   Button "b_Save" at 1074,510 size 72x64; TextOff 'SAVE'; Authorization "Operate"; PictureOff "SetHD"
      on Click: SetBit("DB_MouldEditor_HMI_uData_sStatusBits_xSafeChanges"); "VBStore_tool"('\Storage Card SD')
      Visibility <- "DB_MouldEditor_HMI_uData_sStatusBits_xValueChanged"
   IOField "I/O field_15" at 673,669 size 77x35; Authorization "Operate"; FormatPattern 9999.99
      ProcessValue <- "DB_MouldEditor_HMI_uData_sSelected_sPS_arFlow{3}"
      Visibility <- "DB704_MH_Value_Mixinghead{0}_AmountComponent"
      ObjectEnable <- "DB_MouldEditor_HMI_uData_sSelected_iCalculation"
      Appearance <- "DB_MouldEditor_HMI_uData_sSelected_iCalculation"
      on OnFinishInput: SetBit("DB_MouldEditor_HMI_uData_sStatusBits_xValueChanged")
   IOField "I/O field_16" at 673,703 size 77x35; Authorization "Operate"; FormatPattern 9999.99
      ProcessValue <- "DB_MouldEditor_HMI_uData_sSelected_sPS_arRatio{3}"
      Visibility <- "DB704_MH_Value_Mixinghead{0}_AmountComponent"
      Appearance <- "DB_MouldEditor_HMI_uData_sSelected_sPS_RefComponent"
      ObjectEnable <- "DB_MouldEditor_HMI_uData_sSelected_sPS_RefComponent"
      on OnFinishInput: SetBit("DB_MouldEditor_HMI_uData_sStatusBits_xValueChanged")
   IOField "I/O field_17" at 673,737 size 77x35; Authorization "Operate"; FormatPattern 9999.99
      ProcessValue <- "DB_MouldEditor_HMI_uData_sSelected_sPS_arPressure{3}"
      Visibility <- "DB704_MH_Value_Mixinghead{0}_AmountComponent"
      on OnFinishInput: SetBit("DB_MouldEditor_HMI_uData_sStatusBits_xValueChanged")
   IOField "I/O field_18" at 808,669 size 77x35; Authorization "Operate"; FormatPattern 9999.99
      ProcessValue <- "DB_MouldEditor_HMI_uData_sSelected_sPS_arFlow{4}"
      Visibility <- "DB704_MH_Value_Mixinghead{0}_AmountComponent"
      ObjectEnable <- "DB_MouldEditor_HMI_uData_sSelected_iCalculation"
      Appearance <- "DB_MouldEditor_HMI_uData_sSelected_iCalculation"
      on OnFinishInput: SetBit("DB_MouldEditor_HMI_uData_sStatusBits_xValueChanged")
   IOField "I/O field_19" at 808,703 size 77x35; Authorization "Operate"; FormatPattern 9999.99
      ProcessValue <- "DB_MouldEditor_HMI_uData_sSelected_sPS_arRatio{4}"
      Visibility <- "DB704_MH_Value_Mixinghead{0}_AmountComponent"
      Appearance <- "DB_MouldEditor_HMI_uData_sSelected_sPS_RefComponent"
      ObjectEnable <- "DB_MouldEditor_HMI_uData_sSelected_sPS_RefComponent"
      on OnFinishInput: SetBit("DB_MouldEditor_HMI_uData_sStatusBits_xValueChanged")
   IOField "I/O field_20" at 808,737 size 77x35; Authorization "Operate"; FormatPattern 9999.99
      ProcessValue <- "DB_MouldEditor_HMI_uData_sSelected_sPS_arPressure{4}"
      Visibility <- "DB704_MH_Value_Mixinghead{0}_AmountComponent"
      on OnFinishInput: SetBit("DB_MouldEditor_HMI_uData_sStatusBits_xValueChanged")
   IOField "I/O field_21" at 944,669 size 77x35; Authorization "Operate"; FormatPattern 9999.99
      ProcessValue <- "DB_MouldEditor_HMI_uData_sSelected_sPS_arFlow{5}"
      Visibility <- "DB704_MH_Value_Mixinghead{0}_AmountComponent"
      ObjectEnable <- "DB_MouldEditor_HMI_uData_sSelected_iCalculation"
      Appearance <- "DB_MouldEditor_HMI_uData_sSelected_iCalculation"
      on OnFinishInput: SetBit("DB_MouldEditor_HMI_uData_sStatusBits_xValueChanged")
   IOField "I/O field_22" at 944,703 size 77x35; Authorization "Operate"; FormatPattern 9999.99
      ProcessValue <- "DB_MouldEditor_HMI_uData_sSelected_sPS_arRatio{5}"
      Visibility <- "DB704_MH_Value_Mixinghead{0}_AmountComponent"
      Appearance <- "DB_MouldEditor_HMI_uData_sSelected_sPS_RefComponent"
      ObjectEnable <- "DB_MouldEditor_HMI_uData_sSelected_sPS_RefComponent"
      on OnFinishInput: SetBit("DB_MouldEditor_HMI_uData_sStatusBits_xValueChanged")
   IOField "I/O field_23" at 944,737 size 77x35; Authorization "Operate"; FormatPattern 9999.99
      ProcessValue <- "DB_MouldEditor_HMI_uData_sSelected_sPS_arPressure{5}"
      Visibility <- "DB704_MH_Value_Mixinghead{0}_AmountComponent"
      on OnFinishInput: SetBit("DB_MouldEditor_HMI_uData_sStatusBits_xValueChanged")
   IOField "I/O field_24" at 1080,669 size 77x35; Authorization "Operate"; FormatPattern 9999.99
      ProcessValue <- "DB_MouldEditor_HMI_uData_sSelected_sPS_arFlow{6}"
      Visibility <- "DB704_MH_Value_Mixinghead{0}_AmountComponent"
      ObjectEnable <- "DB_MouldEditor_HMI_uData_sSelected_iCalculation"
      Appearance <- "DB_MouldEditor_HMI_uData_sSelected_iCalculation"
      on OnFinishInput: SetBit("DB_MouldEditor_HMI_uData_sStatusBits_xValueChanged")
   IOField "I/O field_25" at 1080,703 size 77x35; Authorization "Operate"; FormatPattern 9999.99
      ProcessValue <- "DB_MouldEditor_HMI_uData_sSelected_sPS_arRatio{6}"
      Visibility <- "DB704_MH_Value_Mixinghead{0}_AmountComponent"
      Appearance <- "DB_MouldEditor_HMI_uData_sSelected_sPS_RefComponent"
      ObjectEnable <- "DB_MouldEditor_HMI_uData_sSelected_sPS_RefComponent"
      on OnFinishInput: SetBit("DB_MouldEditor_HMI_uData_sStatusBits_xValueChanged")
   IOField "I/O field_26" at 1080,737 size 77x35; Authorization "Operate"; FormatPattern 9999.99
      ProcessValue <- "DB_MouldEditor_HMI_uData_sSelected_sPS_arPressure{6}"
      Visibility <- "DB704_MH_Value_Mixinghead{0}_AmountComponent"
      on OnFinishInput: SetBit("DB_MouldEditor_HMI_uData_sStatusBits_xValueChanged")
   IOField "I/O field_28" at 235,293 size 84x32; Authorization "Operate"; FormatPattern 999
      ProcessValue <- "DB_MouldEditor_HMI_uData_arShotSet{2}_MHNo"
      Visibility <- "DB_MouldEditor_HMI_uData_uTools_PartShot_Amount"
      Appearance <- "DB_MouldEditor_HMI_uData_sSelected_sPS_iPS"
   IOField "Shottime_2" at 318,293 size 150x32; Authorization "Operate"; FormatPattern 99.999
      ProcessValue <- "DB_MouldEditor_HMI_uData_arShotSet{2}_FoamingTime"
      Visibility <- "DB_MouldEditor_HMI_uData_uTools_PartShot_Amount"
      ObjectEnable <- "DB_MouldEditor_HMI_uData_sSelected_iCalculation"
      Appearance <- "DB_MouldEditor_HMI_uData_sSelected_sPS_iPS"
   IOField "totalflow_2" at 467,293 size 144x32; Authorization "Operate"; FormatPattern 9999.99
      ProcessValue <- "DB_MouldEditor_HMI_uData_sCalculatedValues_arTotalFlow{2}"
      Visibility <- "DB_MouldEditor_HMI_uData_uTools_PartShot_Amount"
      ObjectEnable <- "DB_MouldEditor_HMI_uData_sSelected_iCalculation"
      Appearance <- "DB_MouldEditor_HMI_uData_sSelected_sPS_iPS"
   IOField "totalweight_2" at 609,293 size 151x32; Authorization "Operate"; FormatPattern 999.99
      ProcessValue <- "DB_MouldEditor_HMI_uData_arShotSet{2}_PartWeight"
      Visibility <- "DB_MouldEditor_HMI_uData_uTools_PartShot_Amount"
      ObjectEnable <- "DB_MouldEditor_HMI_uData_sSelected_iCalculation"
      Appearance <- "DB_MouldEditor_HMI_uData_sSelected_sPS_iPS"
   IOField "I/O field_32" at 759,293 size 93x32; Authorization "Operate"; FormatPattern 9999
      ProcessValue <- "DB_MouldEditor_HMI_uData_arShotSet{2}_PartCounter"
      Visibility <- "DB_MouldEditor_HMI_uData_uTools_PartShot_Amount"
      Appearance <- "DB_MouldEditor_HMI_uData_sSelected_sPS_iPS"
   IOField "I/O field_34" at 235,327 size 84x32; Authorization "Operate"; FormatPattern 999
      ProcessValue <- "DB_MouldEditor_HMI_uData_arShotSet{3}_MHNo"
      Visibility <- "DB_MouldEditor_HMI_uData_uTools_PartShot_Amount"
      Appearance <- "DB_MouldEditor_HMI_uData_sSelected_sPS_iPS"
   IOField "Shottime_3" at 318,327 size 150x32; Authorization "Operate"; FormatPattern 99.999
      ProcessValue <- "DB_MouldEditor_HMI_uData_arShotSet{3}_FoamingTime"
      Visibility <- "DB_MouldEditor_HMI_uData_uTools_PartShot_Amount"
      ObjectEnable <- "DB_MouldEditor_HMI_uData_sSelected_iCalculation"
      Appearance <- "DB_MouldEditor_HMI_uData_sSelected_sPS_iPS"
   IOField "totalflow_3" at 467,327 size 144x32; Authorization "Operate"; FormatPattern 9999.99
      ProcessValue <- "DB_MouldEditor_HMI_uData_sCalculatedValues_arTotalFlow{3}"
      Visibility <- "DB_MouldEditor_HMI_uData_uTools_PartShot_Amount"
      ObjectEnable <- "DB_MouldEditor_HMI_uData_sSelected_iCalculation"
      Appearance <- "DB_MouldEditor_HMI_uData_sSelected_sPS_iPS"
   IOField "totalweight_3" at 609,327 size 151x32; Authorization "Operate"; FormatPattern 999.99
      ProcessValue <- "DB_MouldEditor_HMI_uData_arShotSet{3}_PartWeight"
      Visibility <- "DB_MouldEditor_HMI_uData_uTools_PartShot_Amount"
      ObjectEnable <- "DB_MouldEditor_HMI_uData_sSelected_iCalculation"
      Appearance <- "DB_MouldEditor_HMI_uData_sSelected_sPS_iPS"
   IOField "I/O field_38" at 759,327 size 93x32; Authorization "Operate"; FormatPattern 9999
      ProcessValue <- "DB_MouldEditor_HMI_uData_arShotSet{3}_PartCounter"
      Visibility <- "DB_MouldEditor_HMI_uData_uTools_PartShot_Amount"
      Appearance <- "DB_MouldEditor_HMI_uData_sSelected_sPS_iPS"
   IOField "I/O field_40" at 235,362 size 84x32; Authorization "Operate"; FormatPattern 999
      ProcessValue <- "DB_MouldEditor_HMI_uData_arShotSet{4}_MHNo"
      Visibility <- "DB_MouldEditor_HMI_uData_uTools_PartShot_Amount"
      Appearance <- "DB_MouldEditor_HMI_uData_sSelected_sPS_iPS"
   IOField "Shottime_4" at 318,362 size 150x32; Authorization "Operate"; FormatPattern 99.999
      ProcessValue <- "DB_MouldEditor_HMI_uData_arShotSet{4}_FoamingTime"
      Visibility <- "DB_MouldEditor_HMI_uData_uTools_PartShot_Amount"
      ObjectEnable <- "DB_MouldEditor_HMI_uData_sSelected_iCalculation"
      Appearance <- "DB_MouldEditor_HMI_uData_sSelected_sPS_iPS"
   IOField "totalflow_4" at 467,362 size 144x32; Authorization "Operate"; FormatPattern 9999.99
      ProcessValue <- "DB_MouldEditor_HMI_uData_sCalculatedValues_arTotalFlow{4}"
      Visibility <- "DB_MouldEditor_HMI_uData_uTools_PartShot_Amount"
      ObjectEnable <- "DB_MouldEditor_HMI_uData_sSelected_iCalculation"
      Appearance <- "DB_MouldEditor_HMI_uData_sSelected_sPS_iPS"
   IOField "totalweight_4" at 609,362 size 151x32; Authorization "Operate"; FormatPattern 999.99
      ProcessValue <- "DB_MouldEditor_HMI_uData_arShotSet{4}_PartWeight"
      Visibility <- "DB_MouldEditor_HMI_uData_uTools_PartShot_Amount"
      ObjectEnable <- "DB_MouldEditor_HMI_uData_sSelected_iCalculation"
      Appearance <- "DB_MouldEditor_HMI_uData_sSelected_sPS_iPS"
   IOField "I/O field_44" at 759,362 size 93x32; Authorization "Operate"; FormatPattern 9999
      ProcessValue <- "DB_MouldEditor_HMI_uData_arShotSet{4}_PartCounter"
      Visibility <- "DB_MouldEditor_HMI_uData_uTools_PartShot_Amount"
      Appearance <- "DB_MouldEditor_HMI_uData_sSelected_sPS_iPS"
   IOField "I/O field_46" at 235,397 size 84x32; Authorization "Operate"; FormatPattern 999
      ProcessValue <- "DB_MouldEditor_HMI_uData_arShotSet{5}_MHNo"
      Visibility <- "DB_MouldEditor_HMI_uData_uTools_PartShot_Amount"
      Appearance <- "DB_MouldEditor_HMI_uData_sSelected_sPS_iPS"
   IOField "Shottime_5" at 318,397 size 150x32; Authorization "Operate"; FormatPattern 99.999
      ProcessValue <- "DB_MouldEditor_HMI_uData_arShotSet{5}_FoamingTime"
      Visibility <- "DB_MouldEditor_HMI_uData_uTools_PartShot_Amount"
      ObjectEnable <- "DB_MouldEditor_HMI_uData_sSelected_iCalculation"
      Appearance <- "DB_MouldEditor_HMI_uData_sSelected_sPS_iPS"
   IOField "totalflow_5" at 467,397 size 144x32; Authorization "Operate"; FormatPattern 9999.99
      ProcessValue <- "DB_MouldEditor_HMI_uData_sCalculatedValues_arTotalFlow{5}"
      Visibility <- "DB_MouldEditor_HMI_uData_uTools_PartShot_Amount"
      ObjectEnable <- "DB_MouldEditor_HMI_uData_sSelected_iCalculation"
      Appearance <- "DB_MouldEditor_HMI_uData_sSelected_sPS_iPS"
   IOField "totalweight_5" at 609,397 size 151x32; Authorization "Operate"; FormatPattern 999.99
      ProcessValue <- "DB_MouldEditor_HMI_uData_arShotSet{5}_PartWeight"
      Visibility <- "DB_MouldEditor_HMI_uData_uTools_PartShot_Amount"
      ObjectEnable <- "DB_MouldEditor_HMI_uData_sSelected_iCalculation"
      Appearance <- "DB_MouldEditor_HMI_uData_sSelected_sPS_iPS"
   IOField "I/O field_50" at 759,397 size 93x32; Authorization "Operate"; FormatPattern 9999
      ProcessValue <- "DB_MouldEditor_HMI_uData_arShotSet{5}_PartCounter"
      Visibility <- "DB_MouldEditor_HMI_uData_uTools_PartShot_Amount"
      Appearance <- "DB_MouldEditor_HMI_uData_sSelected_sPS_iPS"
   IOField "I/O field_52" at 235,432 size 84x32; Authorization "Operate"; FormatPattern 999
      ProcessValue <- "DB_MouldEditor_HMI_uData_arShotSet{6}_MHNo"
      Visibility <- "DB_MouldEditor_HMI_uData_uTools_PartShot_Amount"
      Appearance <- "DB_MouldEditor_HMI_uData_sSelected_sPS_iPS"
   IOField "Shottime_6" at 318,432 size 150x32; Authorization "Operate"; FormatPattern 99.999
      ProcessValue <- "DB_MouldEditor_HMI_uData_arShotSet{6}_FoamingTime"
      Visibility <- "DB_MouldEditor_HMI_uData_uTools_PartShot_Amount"
      ObjectEnable <- "DB_MouldEditor_HMI_uData_sSelected_iCalculation"
      Appearance <- "DB_MouldEditor_HMI_uData_sSelected_sPS_iPS"
   IOField "totalflow_6" at 467,432 size 144x32; Authorization "Operate"; FormatPattern 9999.99
      ProcessValue <- "DB_MouldEditor_HMI_uData_sCalculatedValues_arTotalFlow{6}"
      Visibility <- "DB_MouldEditor_HMI_uData_uTools_PartShot_Amount"
      ObjectEnable <- "DB_MouldEditor_HMI_uData_sSelected_iCalculation"
      Appearance <- "DB_MouldEditor_HMI_uData_sSelected_sPS_iPS"
   IOField "totalweight_6" at 609,432 size 151x32; Authorization "Operate"; FormatPattern 999.99
      ProcessValue <- "DB_MouldEditor_HMI_uData_arShotSet{6}_PartWeight"
      Visibility <- "DB_MouldEditor_HMI_uData_uTools_PartShot_Amount"
      ObjectEnable <- "DB_MouldEditor_HMI_uData_sSelected_iCalculation"
      Appearance <- "DB_MouldEditor_HMI_uData_sSelected_sPS_iPS"
   IOField "I/O field_56" at 759,432 size 93x32; Authorization "Operate"; FormatPattern 9999
      ProcessValue <- "DB_MouldEditor_HMI_uData_arShotSet{6}_PartCounter"
      Visibility <- "DB_MouldEditor_HMI_uData_uTools_PartShot_Amount"
      Appearance <- "DB_MouldEditor_HMI_uData_sSelected_sPS_iPS"
   IOField "I/O field_58" at 235,467 size 84x32; Authorization "Operate"; FormatPattern 999
      ProcessValue <- "DB_MouldEditor_HMI_uData_arShotSet{7}_MHNo"
      Visibility <- "DB_MouldEditor_HMI_uData_uTools_PartShot_Amount"
      Appearance <- "DB_MouldEditor_HMI_uData_sSelected_sPS_iPS"
   IOField "Shottime_7" at 318,467 size 150x32; Authorization "Operate"; FormatPattern 99.999
      ProcessValue <- "DB_MouldEditor_HMI_uData_arShotSet{7}_FoamingTime"
      Visibility <- "DB_MouldEditor_HMI_uData_uTools_PartShot_Amount"
      ObjectEnable <- "DB_MouldEditor_HMI_uData_sSelected_iCalculation"
      Appearance <- "DB_MouldEditor_HMI_uData_sSelected_sPS_iPS"
   IOField "totalflow_7" at 467,467 size 144x32; Authorization "Operate"; FormatPattern 9999.99
      ProcessValue <- "DB_MouldEditor_HMI_uData_sCalculatedValues_arTotalFlow{7}"
      Visibility <- "DB_MouldEditor_HMI_uData_uTools_PartShot_Amount"
      ObjectEnable <- "DB_MouldEditor_HMI_uData_sSelected_iCalculation"
      Appearance <- "DB_MouldEditor_HMI_uData_sSelected_sPS_iPS"
   IOField "totalweight_7" at 609,467 size 151x32; Authorization "Operate"; FormatPattern 999.99
      ProcessValue <- "DB_MouldEditor_HMI_uData_arShotSet{7}_PartWeight"
      Visibility <- "DB_MouldEditor_HMI_uData_uTools_PartShot_Amount"
      ObjectEnable <- "DB_MouldEditor_HMI_uData_sSelected_iCalculation"
      Appearance <- "DB_MouldEditor_HMI_uData_sSelected_sPS_iPS"
   IOField "I/O field_62" at 759,467 size 93x32; Authorization "Operate"; FormatPattern 9999
      ProcessValue <- "DB_MouldEditor_HMI_uData_arShotSet{7}_PartCounter"
      Visibility <- "DB_MouldEditor_HMI_uData_uTools_PartShot_Amount"
      Appearance <- "DB_MouldEditor_HMI_uData_sSelected_sPS_iPS"
   IOField "I/O field_64" at 235,502 size 84x32; Authorization "Operate"; FormatPattern 999
      ProcessValue <- "DB_MouldEditor_HMI_uData_arShotSet{8}_MHNo"
      Visibility <- "DB_MouldEditor_HMI_uData_uTools_PartShot_Amount"
      Appearance <- "DB_MouldEditor_HMI_uData_sSelected_sPS_iPS"
   IOField "Shottime_8" at 318,502 size 150x32; Authorization "Operate"; FormatPattern 99.999
      ProcessValue <- "DB_MouldEditor_HMI_uData_arShotSet{8}_FoamingTime"
      Visibility <- "DB_MouldEditor_HMI_uData_uTools_PartShot_Amount"
      ObjectEnable <- "DB_MouldEditor_HMI_uData_sSelected_iCalculation"
      Appearance <- "DB_MouldEditor_HMI_uData_sSelected_sPS_iPS"
   IOField "totalflow_8" at 467,502 size 144x32; Authorization "Operate"; FormatPattern 9999.99
      ProcessValue <- "DB_MouldEditor_HMI_uData_sCalculatedValues_arTotalFlow{8}"
      Visibility <- "DB_MouldEditor_HMI_uData_uTools_PartShot_Amount"
      ObjectEnable <- "DB_MouldEditor_HMI_uData_sSelected_iCalculation"
      Appearance <- "DB_MouldEditor_HMI_uData_sSelected_sPS_iPS"
   IOField "totalweight_8" at 609,502 size 151x32; Authorization "Operate"; FormatPattern 999.99
      ProcessValue <- "DB_MouldEditor_HMI_uData_arShotSet{8}_PartWeight"
      Visibility <- "DB_MouldEditor_HMI_uData_uTools_PartShot_Amount"
      ObjectEnable <- "DB_MouldEditor_HMI_uData_sSelected_iCalculation"
      Appearance <- "DB_MouldEditor_HMI_uData_sSelected_sPS_iPS"
   IOField "I/O field_68" at 759,502 size 93x32; Authorization "Operate"; FormatPattern 9999
      ProcessValue <- "DB_MouldEditor_HMI_uData_arShotSet{8}_PartCounter"
      Visibility <- "DB_MouldEditor_HMI_uData_uTools_PartShot_Amount"
      Appearance <- "DB_MouldEditor_HMI_uData_sSelected_sPS_iPS"
   Button "b_Shottime" at 368,184 size 48x40; TextOff 'ST'; PictureOff "shottime_1"
      on Click: SetTag("DB_MouldEditor_HMI_uData_sSelected_iCalculation", 0)
   Button "b_TotalFlow" at 514,184 size 48x40; TextOff 'TF'; PictureOff "Actual_Fault_1"
      on Click: SetTag("DB_MouldEditor_HMI_uData_sSelected_iCalculation", 1)
   Button "b_TotalWeight" at 661,184 size 48x40; TextOff 'TW'; PictureOff "Actual_Fault_1"
      on Click: SetTag("DB_MouldEditor_HMI_uData_sSelected_iCalculation", 2)
   Button "b_sub_up" at 103,285 size 40x80; TextOff 'Text'; PictureOff "up arrow"; Authorization "Operate"
      Visibility <- "DB_MouldEditor_HMI_uData_uTools_PartShot_Amount"
      on Click: function_b9b71300("DB_MouldEditor_HMI_uData_uTools_PartShot_Amount", 1)
   Button "b_add_down" at 102,456 size 40x80; TextOff 'Text'; PictureOff "down arrow"; Authorization "Operate"
      Visibility <- "DB_MouldEditor_HMI_uData_uTools_PartShot_Amount"
      on Click: function_dd21b452("DB_MouldEditor_HMI_uData_uTools_PartShot_Amount", 1)
   Button "b_Incress_ToolEditor" at 418,146 size 40x29; TextOff 'Text'; PictureOff "right arrow"
      on Click: function_dd21b452("DB_MouldEditor_HMI_uData_sSelected_iTool", 1)
   Button "check_enabletool" at 874,149 size 40x25; TextOff 'Text'; PictureOff "download"; PictureList "Check_Uncheck"
      ProcessValue <- "DB_MouldEditor_HMI_uData_uTools_EnableTool"
      Visibility <- "DB_MouldEditor_HMI_uData_uTools_PartShot_Amount"
      on Click: InvertBit("DB_MouldEditor_HMI_uData_uTools_EnableTool")
   Button "check_Service_1" at 870,262 size 40x25; TextOff 'Text'; PictureOff "download"; PictureList "Check_Uncheck"
      Visibility <- "DB_MouldEditor_HMI_uData_uTools_PartShot_Amount"
      ProcessValue <- "DB_MouldEditor_HMI_uData_arShotSet{1}_PartShotDisable"
      on Click: InvertBit("DB_MouldEditor_HMI_uData_arShotSet{1}_PartShotDisable")
   Button "check_Service_2" at 870,297 size 40x25; TextOff 'Text'; PictureOff "download"; PictureList "Check_Uncheck"
      Visibility <- "DB_MouldEditor_HMI_uData_uTools_PartShot_Amount"
      ProcessValue <- "DB_MouldEditor_HMI_uData_arShotSet{2}_PartShotDisable"
      on Click: InvertBit("DB_MouldEditor_HMI_uData_arShotSet{2}_PartShotDisable")
   Button "check_Service_3" at 870,331 size 40x25; TextOff 'Text'; PictureOff "download"; PictureList "Check_Uncheck"
      Visibility <- "DB_MouldEditor_HMI_uData_uTools_PartShot_Amount"
      ProcessValue <- "DB_MouldEditor_HMI_uData_arShotSet{3}_PartShotDisable"
      on Click: InvertBit("DB_MouldEditor_HMI_uData_arShotSet{3}_PartShotDisable")
   Button "check_Service_4" at 870,366 size 40x25; TextOff 'Text'; PictureOff "download"; PictureList "Check_Uncheck"
      Visibility <- "DB_MouldEditor_HMI_uData_uTools_PartShot_Amount"
      ProcessValue <- "DB_MouldEditor_HMI_uData_arShotSet{4}_PartShotDisable"
      on Click: InvertBit("DB_MouldEditor_HMI_uData_arShotSet{4}_PartShotDisable")
   Button "check_Service_5" at 870,401 size 40x25; TextOff 'Text'; PictureOff "download"; PictureList "Check_Uncheck"
      Visibility <- "DB_MouldEditor_HMI_uData_uTools_PartShot_Amount"
      ProcessValue <- "DB_MouldEditor_HMI_uData_arShotSet{5}_PartShotDisable"
      on Click: InvertBit("DB_MouldEditor_HMI_uData_arShotSet{5}_PartShotDisable")
   Button "check_Service_6" at 870,436 size 40x25; TextOff 'Text'; PictureOff "download"; PictureList "Check_Uncheck"
      Visibility <- "DB_MouldEditor_HMI_uData_uTools_PartShot_Amount"
      ProcessValue <- "DB_MouldEditor_HMI_uData_arShotSet{6}_PartShotDisable"
      on Click: InvertBit("DB_MouldEditor_HMI_uData_arShotSet{6}_PartShotDisable")
   Button "check_Service_7" at 870,471 size 40x25; TextOff 'Text'; PictureOff "download"; PictureList "Check_Uncheck"
      Visibility <- "DB_MouldEditor_HMI_uData_uTools_PartShot_Amount"
      ProcessValue <- "DB_MouldEditor_HMI_uData_arShotSet{7}_PartShotDisable"
      on Click: InvertBit("DB_MouldEditor_HMI_uData_arShotSet{7}_PartShotDisable")
   Button "check_Service_8" at 870,506 size 40x25; TextOff 'Text'; PictureOff "download"; PictureList "Check_Uncheck"
      Visibility <- "DB_MouldEditor_HMI_uData_uTools_PartShot_Amount"
      ProcessValue <- "DB_MouldEditor_HMI_uData_arShotSet{8}_PartShotDisable"
      on Click: InvertBit("DB_MouldEditor_HMI_uData_arShotSet{8}_PartShotDisable")
   Button "check_CP_1" at 941,262 size 40x25; TextOff 'Text'; PictureOff "download"; PictureList "Check_Uncheck"
      ProcessValue <- "DB_MouldEditor_HMI_uData_arShotSet{1}_CPMoveAfterShot"
      Visibility <- "DB_MouldEditor_HMI_uData_uTools_PartShot_Amount"
      on Click: InvertBit("DB_MouldEditor_HMI_uData_arShotSet{1}_CPMoveAfterShot")
   Button "check_CP_2" at 941,297 size 40x25; TextOff 'Text'; PictureOff "download"; PictureList "Check_Uncheck"
      ProcessValue <- "DB_MouldEditor_HMI_uData_arShotSet{2}_CPMoveAfterShot"
      Visibility <- "DB_MouldEditor_HMI_uData_uTools_PartShot_Amount"
      on Click: InvertBit("DB_MouldEditor_HMI_uData_arShotSet{2}_CPMoveAfterShot")
   Button "check_CP_3" at 941,331 size 40x25; TextOff 'Text'; PictureOff "download"; PictureList "Check_Uncheck"
      ProcessValue <- "DB_MouldEditor_HMI_uData_arShotSet{3}_CPMoveAfterShot"
      Visibility <- "DB_MouldEditor_HMI_uData_uTools_PartShot_Amount"
      on Click: InvertBit("DB_MouldEditor_HMI_uData_arShotSet{3}_CPMoveAfterShot")
   Button "check_CP_4" at 941,366 size 40x25; TextOff 'Text'; PictureOff "download"; PictureList "Check_Uncheck"
      ProcessValue <- "DB_MouldEditor_HMI_uData_arShotSet{4}_CPMoveAfterShot"
      Visibility <- "DB_MouldEditor_HMI_uData_uTools_PartShot_Amount"
      on Click: InvertBit("DB_MouldEditor_HMI_uData_arShotSet{4}_CPMoveAfterShot")
   Button "check_CP_5" at 941,401 size 40x25; TextOff 'Text'; PictureOff "download"; PictureList "Check_Uncheck"
      ProcessValue <- "DB_MouldEditor_HMI_uData_arShotSet{5}_CPMoveAfterShot"
      Visibility <- "DB_MouldEditor_HMI_uData_uTools_PartShot_Amount"
      on Click: InvertBit("DB_MouldEditor_HMI_uData_arShotSet{5}_CPMoveAfterShot")
   Button "check_CP_6" at 941,436 size 40x25; TextOff 'Text'; PictureOff "download"; PictureList "Check_Uncheck"
      ProcessValue <- "DB_MouldEditor_HMI_uData_arShotSet{6}_CPMoveAfterShot"
      Visibility <- "DB_MouldEditor_HMI_uData_uTools_PartShot_Amount"
      on Click: InvertBit("DB_MouldEditor_HMI_uData_arShotSet{6}_CPMoveAfterShot")
   Button "check_CP_7" at 941,471 size 40x25; TextOff 'Text'; PictureOff "download"; PictureList "Check_Uncheck"
      ProcessValue <- "DB_MouldEditor_HMI_uData_arShotSet{7}_CPMoveAfterShot"
      Visibility <- "DB_MouldEditor_HMI_uData_uTools_PartShot_Amount"
      on Click: InvertBit("DB_MouldEditor_HMI_uData_arShotSet{7}_CPMoveAfterShot")
   Button "check_CP_8" at 941,506 size 40x25; TextOff 'Text'; PictureOff "download"; PictureList "Check_Uncheck"
      ProcessValue <- "DB_MouldEditor_HMI_uData_arShotSet{8}_CPMoveAfterShot"
      Visibility <- "DB_MouldEditor_HMI_uData_uTools_PartShot_Amount"
      on Click: InvertBit("DB_MouldEditor_HMI_uData_arShotSet{8}_CPMoveAfterShot")
   Button "check_blowingaftershot_1" at 1007,262 size 40x25; TextOff 'Text'; PictureOff "download"; PictureList "Check_Uncheck"
      Visibility <- "DB_MouldEditor_HMI_uData_uTools_PartShot_Amount"
      ProcessValue <- "DB_MouldEditor_HMI_uData_arShotSet{1}_PurgeMHAfterShot"
      on Click: InvertBit("DB_MouldEditor_HMI_uData_arShotSet{1}_PurgeMHAfterShot")
   Button "check_blowingaftershot_2" at 1007,297 size 40x25; TextOff 'Text'; PictureOff "download"; PictureList "Check_Uncheck"
      Visibility <- "DB_MouldEditor_HMI_uData_uTools_PartShot_Amount"
      ProcessValue <- "DB_MouldEditor_HMI_uData_arShotSet{2}_PurgeMHAfterShot"
      on Click: InvertBit("DB_MouldEditor_HMI_uData_arShotSet{2}_PurgeMHAfterShot")
   Button "check_blowingaftershot_3" at 1007,331 size 40x25; TextOff 'Text'; PictureOff "download"; PictureList "Check_Uncheck"
      Visibility <- "DB_MouldEditor_HMI_uData_uTools_PartShot_Amount"
      ProcessValue <- "DB_MouldEditor_HMI_uData_arShotSet{3}_PurgeMHAfterShot"
      on Click: InvertBit("DB_MouldEditor_HMI_uData_arShotSet{3}_PurgeMHAfterShot")
   Button "check_blowingaftershot_4" at 1007,366 size 40x25; TextOff 'Text'; PictureOff "download"; PictureList "Check_Uncheck"
      Visibility <- "DB_MouldEditor_HMI_uData_uTools_PartShot_Amount"
      ProcessValue <- "DB_MouldEditor_HMI_uData_arShotSet{4}_PurgeMHAfterShot"
      on Click: InvertBit("DB_MouldEditor_HMI_uData_arShotSet{4}_PurgeMHAfterShot")
   Button "check_blowingaftershot_5" at 1007,401 size 40x25; TextOff 'Text'; PictureOff "download"; PictureList "Check_Uncheck"
      Visibility <- "DB_MouldEditor_HMI_uData_uTools_PartShot_Amount"
      ProcessValue <- "DB_MouldEditor_HMI_uData_arShotSet{5}_PurgeMHAfterShot"
      on Click: InvertBit("DB_MouldEditor_HMI_uData_arShotSet{5}_PurgeMHAfterShot")
   Button "check_blowingaftershot_6" at 1007,436 size 40x25; TextOff 'Text'; PictureOff "download"; PictureList "Check_Uncheck"
      Visibility <- "DB_MouldEditor_HMI_uData_uTools_PartShot_Amount"
      ProcessValue <- "DB_MouldEditor_HMI_uData_arShotSet{6}_PurgeMHAfterShot"
      on Click: InvertBit("DB_MouldEditor_HMI_uData_arShotSet{6}_PurgeMHAfterShot")
   Button "check_blowingaftershot_7" at 1007,471 size 40x25; TextOff 'Text'; PictureOff "download"; PictureList "Check_Uncheck"
      Visibility <- "DB_MouldEditor_HMI_uData_uTools_PartShot_Amount"
      ProcessValue <- "DB_MouldEditor_HMI_uData_arShotSet{7}_PurgeMHAfterShot"
      on Click: InvertBit("DB_MouldEditor_HMI_uData_arShotSet{7}_PurgeMHAfterShot")
   Button "check_blowingaftershot_8" at 1007,506 size 40x25; TextOff 'Text'; PictureOff "download"; PictureList "Check_Uncheck"
      Visibility <- "DB_MouldEditor_HMI_uData_uTools_PartShot_Amount"
      ProcessValue <- "DB_MouldEditor_HMI_uData_arShotSet{8}_PurgeMHAfterShot"
      on Click: InvertBit("DB_MouldEditor_HMI_uData_arShotSet{8}_PurgeMHAfterShot")
   Button "b_Import" at 997,92 size 80x56; TextOff 'Import USB'; Authorization "User administration"; PictureOff "fromUSB"
      on Click: function_f12b67b1('*.csv', '\Storage Card USB', 1, 1, 1, 0, "ImportDataFrom_USB", "ImportDataFrom_USB_stat"); "ReadDataFromUSB"()
      Visibility <- "NavUserChange"
   Button "b_Export" at 1085,92 size 80x56; TextOff 'Import SD'; Authorization "User administration"; PictureOff "fromSD"
      on Click: function_f12b67b1('*.csv', '\Storage Card SD\Tools', 1, 1, 1, 0, "ImportDataFrom_SD", "ImportDataFrom_SD_stat"); "ReadDataFromSD"()
      Visibility <- "NavUserChange"
   Button "Button_9" at 148,258 size 86x32; TextOff '1.'
      Visibility <- "DB_MouldEditor_HMI_uData_uTools_PartShot_Amount"
      Appearance <- "DB_MouldEditor_HMI_uData_sSelected_sPS_iPS"
   Button "Button_10" at 148,293 size 86x32; TextOff '2.'
      Visibility <- "DB_MouldEditor_HMI_uData_uTools_PartShot_Amount"
      Appearance <- "DB_MouldEditor_HMI_uData_sSelected_sPS_iPS"
   Button "Button_11" at 148,327 size 86x32; TextOff '3.'
      Visibility <- "DB_MouldEditor_HMI_uData_uTools_PartShot_Amount"
      Appearance <- "DB_MouldEditor_HMI_uData_sSelected_sPS_iPS"
   Button "Button_12" at 148,362 size 86x32; TextOff '4.'
      Visibility <- "DB_MouldEditor_HMI_uData_uTools_PartShot_Amount"
      Appearance <- "DB_MouldEditor_HMI_uData_sSelected_sPS_iPS"
   Button "Button_13" at 148,397 size 86x32; TextOff '5.'
      Visibility <- "DB_MouldEditor_HMI_uData_uTools_PartShot_Amount"
      Appearance <- "DB_MouldEditor_HMI_uData_sSelected_sPS_iPS"
   Button "Button_14" at 148,432 size 86x32; TextOff '6.'
      Visibility <- "DB_MouldEditor_HMI_uData_uTools_PartShot_Amount"
      Appearance <- "DB_MouldEditor_HMI_uData_sSelected_sPS_iPS"
   Button "Button_15" at 148,467 size 86x32; TextOff '7.'
      Visibility <- "DB_MouldEditor_HMI_uData_uTools_PartShot_Amount"
      Appearance <- "DB_MouldEditor_HMI_uData_sSelected_sPS_iPS"
   Button "Button_16" at 148,502 size 86x32; TextOff '8.'
      Visibility <- "DB_MouldEditor_HMI_uData_uTools_PartShot_Amount"
      Appearance <- "DB_MouldEditor_HMI_uData_sSelected_sPS_iPS"
   Button "b_Decress_Tool_Editor" at 310,146 size 40x29; TextOff 'Text'; PictureOff "left arrow"
      on Click: function_b9b71300("DB_MouldEditor_HMI_uData_sSelected_iTool", 1)
      Visibility <- "DB_MouldEditor_HMI_uData_sSelected_iTool"
   Button "b_SetHD" at 1075,431 size 72x64; TextOff 'SetHD'; Authorization "Operate"; PictureOff "Save_Icon"
      on Click: SetBit("InterfaceVisu_SetHDValue")
      Visibility <- "DB_MouldEditor_HMI_uData_sStatusBits_xValueChanged"
      Appearance <- "InterfaceVisu_HPValuesSet"
   TextField "Text field_14" at 994,201 size 66x58; Text 'Blowing After Shot'
      Visibility <- "DB704_MH_Value_Mixinghead{0}_WithInerting"
   Circle "Circle_1" at 1094,446 size 34x34
      Visibility <- "DB_MouldEditor_HMI_uData_sStatusBits_xValueChanged"
   Circle "Circle_2" at 1085,437 size 52x52
      Visibility <- "DB_MouldEditor_HMI_uData_sStatusBits_xValueChanged"
   Button "b_SetHD_1" at 1075,431 size 72x64; TextOff 'SetHD'; Authorization "Operate"; PictureOff "Save_Icon"
      on Click: SetBit("InterfaceVisu_SetHDValue")
      Visibility <- "DB_MouldEditor_HMI_uData_sStatusBits_xValueChanged"
      Appearance <- "InterfaceVisu_SetHDValue"
   Button "Button_2" at 350,627 size 130x32; TextOff 'Text'; TextList "Pump_Name"
      ObjectEnable <- "Activate_Deactivate"
      on Press: SetTag("DB_MouldEditor_HMI_uData_sSelected_sPS_RefComponent", 1)
      Appearance <- "DB_MouldEditor_HMI_uData_sSelected_sPS_RefComponent"
      ProcessValue <- "DB704_MH_Value_Mixinghead{0}_MH_Connection{1}_Pump_No"
      Visibility <- "DB704_MH_Value_Mixinghead{0}_AmountComponent"
   Button "Button_4" at 486,627 size 130x32; TextOff 'Text'; TextList "Pump_Name"
      ObjectEnable <- "Activate_Deactivate"
      on Press: SetTag("DB_MouldEditor_HMI_uData_sSelected_sPS_RefComponent", 2)
      Appearance <- "DB_MouldEditor_HMI_uData_sSelected_sPS_RefComponent"
      ProcessValue <- "DB704_MH_Value_Mixinghead{0}_MH_Connection{2}_Pump_No"
      Visibility <- "DB704_MH_Value_Mixinghead{0}_AmountComponent"
   Button "Button_5" at 620,627 size 130x32; TextOff 'Text'; TextList "Pump_Name"
      ObjectEnable <- "Activate_Deactivate"
      on Press: SetTag("DB_MouldEditor_HMI_uData_sSelected_sPS_RefComponent", 3)
      Appearance <- "DB_MouldEditor_HMI_uData_sSelected_sPS_RefComponent"
      ProcessValue <- "DB704_MH_Value_Mixinghead{0}_MH_Connection{3}_Pump_No"
      Visibility <- "DB704_MH_Value_Mixinghead{0}_AmountComponent"
   Button "Button_6" at 755,627 size 130x32; TextOff 'Text'; TextList "Pump_Name"
      ObjectEnable <- "Activate_Deactivate"
      on Press: SetTag("DB_MouldEditor_HMI_uData_sSelected_sPS_RefComponent", 4)
      Appearance <- "DB_MouldEditor_HMI_uData_sSelected_sPS_RefComponent"
      ProcessValue <- "DB704_MH_Value_Mixinghead{0}_MH_Connection{4}_Pump_No"
      Visibility <- "DB704_MH_Value_Mixinghead{0}_AmountComponent"
   Button "Button_7" at 891,627 size 130x32; TextOff 'Text'; TextList "Pump_Name"
      ObjectEnable <- "Activate_Deactivate"
      on Press: SetTag("DB_MouldEditor_HMI_uData_sSelected_sPS_RefComponent", 5)
      Appearance <- "DB_MouldEditor_HMI_uData_sSelected_sPS_RefComponent"
      ProcessValue <- "DB704_MH_Value_Mixinghead{0}_MH_Connection{5}_Pump_No"
      Visibility <- "DB704_MH_Value_Mixinghead{0}_AmountComponent"
   Button "Button_8" at 1027,627 size 130x32; TextOff 'Text'; TextList "Pump_Name"
      ObjectEnable <- "Activate_Deactivate"
      on Press: SetTag("DB_MouldEditor_HMI_uData_sSelected_sPS_RefComponent", 6)
      Appearance <- "DB_MouldEditor_HMI_uData_sSelected_sPS_RefComponent"
      ProcessValue <- "DB704_MH_Value_Mixinghead{0}_MH_Connection{6}_Pump_No"
      Visibility <- "DB704_MH_Value_Mixinghead{0}_AmountComponent"
   IOField "Shottime_9" at 318,258 size 150x32; Authorization "Operate"; FormatPattern 99.999
      ProcessValue <- "DB_MouldEditor_HMI_uData_arShotSet{1}_FoamingTime"
      Visibility <- "DB_MouldEditor_HMI_uData_sColumn_iShotTime"
   IOField "Shottime_10" at 318,293 size 150x32; Authorization "Operate"; FormatPattern 99.999
      ProcessValue <- "DB_MouldEditor_HMI_uData_arShotSet{2}_FoamingTime"
      Visibility <- "DB_MouldEditor_HMI_uData_sColumn_iShotTime"
   IOField "Shottime_11" at 318,327 size 150x32; Authorization "Operate"; FormatPattern 99.999
      ProcessValue <- "DB_MouldEditor_HMI_uData_arShotSet{3}_FoamingTime"
      Visibility <- "DB_MouldEditor_HMI_uData_sColumn_iShotTime"
   IOField "Shottime_12" at 318,362 size 150x32; Authorization "Operate"; FormatPattern 99.999
      ProcessValue <- "DB_MouldEditor_HMI_uData_arShotSet{4}_FoamingTime"
      Visibility <- "DB_MouldEditor_HMI_uData_sColumn_iShotTime"
   IOField "Shottime_13" at 318,397 size 150x32; Authorization "Operate"; FormatPattern 99.999
      ProcessValue <- "DB_MouldEditor_HMI_uData_arShotSet{5}_FoamingTime"
      Visibility <- "DB_MouldEditor_HMI_uData_sColumn_iShotTime"
   IOField "Shottime_14" at 318,432 size 150x32; Authorization "Operate"; FormatPattern 99.999
      ProcessValue <- "DB_MouldEditor_HMI_uData_arShotSet{6}_FoamingTime"
      Visibility <- "DB_MouldEditor_HMI_uData_sColumn_iShotTime"
   IOField "Shottime_15" at 318,467 size 150x32; Authorization "Operate"; FormatPattern 99.999
      ProcessValue <- "DB_MouldEditor_HMI_uData_arShotSet{7}_FoamingTime"
      Visibility <- "DB_MouldEditor_HMI_uData_sColumn_iShotTime"
   IOField "Shottime_16" at 318,502 size 150x32; Authorization "Operate"; FormatPattern 99.999
      ProcessValue <- "DB_MouldEditor_HMI_uData_arShotSet{8}_FoamingTime"
      Visibility <- "DB_MouldEditor_HMI_uData_sColumn_iShotTime"
   IOField "totalflow_9" at 467,258 size 144x32; Authorization "Operate"; FormatPattern 9999.99
      ProcessValue <- "DB_MouldEditor_HMI_uData_sCalculatedValues_arTotalFlow{1}"
      Visibility <- "DB_MouldEditor_HMI_uData_sColumn_iTotalFlow"
   IOField "totalflow_10" at 467,293 size 144x32; Authorization "Operate"; FormatPattern 9999.99
      ProcessValue <- "DB_MouldEditor_HMI_uData_sCalculatedValues_arTotalFlow{2}"
      Visibility <- "DB_MouldEditor_HMI_uData_sColumn_iTotalFlow"
   IOField "totalflow_11" at 467,327 size 144x32; Authorization "Operate"; FormatPattern 9999.99
      ProcessValue <- "DB_MouldEditor_HMI_uData_sCalculatedValues_arTotalFlow{3}"
      Visibility <- "DB_MouldEditor_HMI_uData_sColumn_iTotalFlow"
   IOField "totalflow_12" at 467,362 size 144x32; Authorization "Operate"; FormatPattern 9999.99
      ProcessValue <- "DB_MouldEditor_HMI_uData_sCalculatedValues_arTotalFlow{4}"
      Visibility <- "DB_MouldEditor_HMI_uData_sColumn_iTotalFlow"
   IOField "totalflow_13" at 467,397 size 144x32; Authorization "Operate"; FormatPattern 9999.99
      ProcessValue <- "DB_MouldEditor_HMI_uData_sCalculatedValues_arTotalFlow{5}"
      Visibility <- "DB_MouldEditor_HMI_uData_sColumn_iTotalFlow"
   IOField "totalflow_14" at 467,432 size 144x32; Authorization "Operate"; FormatPattern 9999.99
      ProcessValue <- "DB_MouldEditor_HMI_uData_sCalculatedValues_arTotalFlow{6}"
      Visibility <- "DB_MouldEditor_HMI_uData_sColumn_iTotalFlow"
   IOField "totalflow_15" at 467,467 size 144x32; Authorization "Operate"; FormatPattern 9999.99
      ProcessValue <- "DB_MouldEditor_HMI_uData_sCalculatedValues_arTotalFlow{7}"
      Visibility <- "DB_MouldEditor_HMI_uData_sColumn_iTotalFlow"
   IOField "totalflow_16" at 467,502 size 144x32; Authorization "Operate"; FormatPattern 9999.99
      ProcessValue <- "DB_MouldEditor_HMI_uData_sCalculatedValues_arTotalFlow{8}"
      Visibility <- "DB_MouldEditor_HMI_uData_sColumn_iTotalFlow"
   IOField "totalweight_9" at 609,258 size 151x32; Authorization "Operate"; FormatPattern 999.99
      ProcessValue <- "DB_MouldEditor_HMI_uData_arShotSet{1}_PartWeight"
      Visibility <- "DB_MouldEditor_HMI_uData_sColumn_iTotalWeight"
   IOField "totalweight_10" at 609,293 size 151x32; Authorization "Operate"; FormatPattern 999.99
      ProcessValue <- "DB_MouldEditor_HMI_uData_arShotSet{2}_PartWeight"
      Visibility <- "DB_MouldEditor_HMI_uData_sColumn_iTotalWeight"
   IOField "totalweight_11" at 609,327 size 151x32; Authorization "Operate"; FormatPattern 999.99
      ProcessValue <- "DB_MouldEditor_HMI_uData_arShotSet{3}_PartWeight"
      Visibility <- "DB_MouldEditor_HMI_uData_sColumn_iTotalWeight"
   IOField "totalweight_12" at 609,362 size 151x32; Authorization "Operate"; FormatPattern 999.99
      ProcessValue <- "DB_MouldEditor_HMI_uData_arShotSet{4}_PartWeight"
      Visibility <- "DB_MouldEditor_HMI_uData_sColumn_iTotalWeight"
   IOField "totalweight_13" at 609,397 size 151x32; Authorization "Operate"; FormatPattern 999.99
      ProcessValue <- "DB_MouldEditor_HMI_uData_arShotSet{5}_PartWeight"
      Visibility <- "DB_MouldEditor_HMI_uData_sColumn_iTotalWeight"
   IOField "totalweight_14" at 609,432 size 151x32; Authorization "Operate"; FormatPattern 999.99
      ProcessValue <- "DB_MouldEditor_HMI_uData_arShotSet{6}_PartWeight"
      Visibility <- "DB_MouldEditor_HMI_uData_sColumn_iTotalWeight"
   IOField "totalweight_15" at 609,467 size 151x32; Authorization "Operate"; FormatPattern 999.99
      ProcessValue <- "DB_MouldEditor_HMI_uData_arShotSet{7}_PartWeight"
      Visibility <- "DB_MouldEditor_HMI_uData_sColumn_iTotalWeight"
   IOField "totalweight_16" at 609,502 size 151x32; Authorization "Operate"; FormatPattern 999.99
      ProcessValue <- "DB_MouldEditor_HMI_uData_arShotSet{8}_PartWeight"
      Visibility <- "DB_MouldEditor_HMI_uData_sColumn_iTotalWeight"
   Rectangle "Rectangle_22" at 994,159 size 78x376
      Visibility <- "DB704_MH_Value_Mixinghead{0}_WithInerting"
   Button "b_ToolAlloc" at 1071,243 size 80x80; TextOff 'Text'
      Visibility <- "DB_MouldEditor_HMI_uData_sStatusBits_xValueChanged"
      on Click: function_efd93a16("Save", 446, 387, -1, -1, 1)
   Button "b_Part_Counter" at 1074,352 size 73x65; TextOff 'Text'
      Visibility <- "DB_MouldEditor_HMI_uData_sStatusBits_xValueChanged"
      on Click: function_efd93a16("Save", 446, 387, -1, -1, 1)
   Rectangle "Rectangle_1" at 1065,188 size 97x83
      Visibility <- "DB_MouldEditor_HMI_uData_uTools_PartShot_Amount"
   Rectangle "Rectangle_4" at 103,578 size 1061x205
      Visibility <- "DB_MouldEditor_HMI_uData_uTools_PartShot_Amount"
   Rectangle "Rectangle_6" at 1065,420 size 97x83
      Visibility <- "DB_MouldEditor_HMI_uData_uTools_PartShot_Amount"
   Button "Button_42" at 146,254 size 919x40; TextOff 'Text'
      on Click: SetTag("DB_MouldEditor_HMI_uData_sSelected_sPS_iPS", 1)
      Visibility <- "DB_MouldEditor_HMI_uData_sSelected_sPS_iPS"
      ObjectEnable <- "DB_MouldEditor_HMI_uData_uTools_PartShot_Amount"
   Button "Button_43" at 146,289 size 919x40; TextOff 'Text'
      Visibility <- "DB_MouldEditor_HMI_uData_sSelected_sPS_iPS"
      ObjectEnable <- "DB_MouldEditor_HMI_uData_uTools_PartShot_Amount"
      Appearance <- "DB_MouldEditor_HMI_uData_sSelected_sPS_iPS"
      on Click: SetTag("DB_MouldEditor_HMI_uData_sSelected_sPS_iPS", 2)
   Button "Button_44" at 146,323 size 919x40; TextOff 'Text'
      Visibility <- "DB_MouldEditor_HMI_uData_sSelected_sPS_iPS"
      ObjectEnable <- "DB_MouldEditor_HMI_uData_uTools_PartShot_Amount"
      Appearance <- "DB_MouldEditor_HMI_uData_sSelected_sPS_iPS"
      on Click: SetTag("DB_MouldEditor_HMI_uData_sSelected_sPS_iPS", 3)
   Button "Button_45" at 146,358 size 919x40; TextOff 'Text'
      Visibility <- "DB_MouldEditor_HMI_uData_sSelected_sPS_iPS"
      ObjectEnable <- "DB_MouldEditor_HMI_uData_uTools_PartShot_Amount"
      Appearance <- "DB_MouldEditor_HMI_uData_sSelected_sPS_iPS"
      on Click: SetTag("DB_MouldEditor_HMI_uData_sSelected_sPS_iPS", 4)
   Button "Button_46" at 146,393 size 919x40; TextOff 'Text'
      Visibility <- "DB_MouldEditor_HMI_uData_sSelected_sPS_iPS"
      ObjectEnable <- "DB_MouldEditor_HMI_uData_uTools_PartShot_Amount"
      Appearance <- "DB_MouldEditor_HMI_uData_sSelected_sPS_iPS"
      on Click: SetTag("DB_MouldEditor_HMI_uData_sSelected_sPS_iPS", 5)
   Button "Button_47" at 146,428 size 919x40; TextOff 'Text'
      Visibility <- "DB_MouldEditor_HMI_uData_sSelected_sPS_iPS"
      ObjectEnable <- "DB_MouldEditor_HMI_uData_uTools_PartShot_Amount"
      Appearance <- "DB_MouldEditor_HMI_uData_sSelected_sPS_iPS"
      on Click: SetTag("DB_MouldEditor_HMI_uData_sSelected_sPS_iPS", 6)
   Button "Button_48" at 146,463 size 919x40; TextOff 'Text'
      Visibility <- "DB_MouldEditor_HMI_uData_sSelected_sPS_iPS"
      ObjectEnable <- "DB_MouldEditor_HMI_uData_uTools_PartShot_Amount"
      Appearance <- "DB_MouldEditor_HMI_uData_sSelected_sPS_iPS"
      on Click: SetTag("DB_MouldEditor_HMI_uData_sSelected_sPS_iPS", 7)
   Button "Button_49" at 146,500 size 919x40; TextOff 'Text'
      Visibility <- "DB_MouldEditor_HMI_uData_sSelected_sPS_iPS"
      ObjectEnable <- "DB_MouldEditor_HMI_uData_uTools_PartShot_Amount"
      Appearance <- "DB_MouldEditor_HMI_uData_sSelected_sPS_iPS"
      on Click: SetTag("DB_MouldEditor_HMI_uData_sSelected_sPS_iPS", 8)
   Button "Template_Button_14" at 410,141 size 54x39; TextOff 'Text'
      on Click: function_efd93a16("Save", 446, 387, -1, -1, 1)
      Visibility <- "DB_MouldEditor_HMI_uData_sStatusBits_xValueChanged"
      ObjectEnable <- "PopUp_Restrict"
   Button "Template_Button_1" at 298,141 size 54x39; TextOff 'Text'
      on Click: function_efd93a16("Save", 446, 387, -1, -1, 1)
      Visibility <- "DB_MouldEditor_HMI_uData_sStatusBits_xValueChanged"
      ObjectEnable <- "PopUp_Restrict"

